       IF #INO_tTrack.rgtTrackMachine[#IN_dMachineIndex].tUserData.dGetDownstreamIndex >= 0 THEN
           #AUX_xValidDwCap := TRUE;
           #OS_xNewCapDw := TRUE;            
           #AUX_dDwCapIndex := #INO_tTrack.rgtTrackMachine[#IN_dMachineIndex].tUserData.dGetDownstreamIndex;
       ELSE
           #AUX_xValidDwCap := FALSE;
           #OS_xNewCapDw := FALSE;            
           #AUX_dDwCapIndex := 0;
       END_IF;

       #INO_tTrack.rgtTrackMachine[#IN_dMachineIndex].tUserData.xGetPosReach := FALSE;

   END_IF;
END_REGION

REGION Network 6: ####_HMI_LOGICS_####
END_REGION

REGION Network 7 (SCL): List of HMI logics
   REGION UpdateDistanceSnaproll

   IF #tHMW.xUpdateDistSnap THEN
       #tHMW.xUpdateDistSnap := FALSE;

       #tHMR.dDistanceFromSnaproll_cmm := #tHMW.dDistanceFromSnaproll_cmm;

   END_IF;

   END_REGION
END_REGION

REGION Network 8: ####_ALARMS_####
END_REGION

REGION Network 9 (SCL): Reset alarms
   IF #IN_xResetAlarms THEN

       #TMP_dwValue := 0;

       SCATTER(IN:=#TMP_dwValue,
               OUT=>#tALM.tF);

       SCATTER(IN:=#TMP_dwValue,
               OUT=>#tALM.tS);

       SCATTER(IN:=#TMP_dwValue,
               OUT=>#tALM.tW);

   END_IF;
END_REGION

REGION Network 10: ####_STATUSES_####
END_REGION

REGION Network 11 (SCL): Calculate alarm statuses
   GATHER(IN:=#tALM.tS,
          OUT=>#TMP_dwValue);

   IF #TMP_dwValue <> 0 THEN
       #ST_xStoppingFaults := TRUE;
   ELSE
       #ST_xStoppingFaults := FALSE;
   END_IF;

   GATHER(IN:=#tALM.tF,
          OUT=>#TMP_dwValue);

   IF #TMP_dwValue <> 0 THEN
       #ST_xFaults := TRUE;
   ELSE
       #ST_xFaults := FALSE;
   END_IF;

   GATHER(IN:=#tALM.tW,
          OUT=>#TMP_dwValue);

   IF #TMP_dwValue <> 0 THEN
       #ST_xWarnings := TRUE;
   ELSE
       #ST_xWarnings := FALSE;
   END_IF;
END_REGION

REGION Network 12 (SCL): Glass break calculation
   #INO_tRibbon.rgtGlassBreakRequest[#IN_dGlassBreakMachineIndex].IN_dDistanceSnaproll_cmm := #tHMR.dDistanceFromSnaproll_cmm;
   #INO_tRibbon.rgtGlassBreakRequest[#IN_dGlassBreakMachineIndex].IN_dDownstreamOffset_cmm := #CONST_DBREAKDOWNOFF_CMM;
   #INO_tRibbon.rgtGlassBreakRequest[#IN_dGlassBreakMachineIndex].IN_dUpstreamOffset_cmm := #CONST_DBREAKUPOFF_CMM;

   IF #INO_tRibbon.rgtGlassBreakRequest[#IN_dGlassBreakMachineIndex].OUT_xDataReady THEN
       #ST_xGlassBreak := #INO_tRibbon.rgtGlassBreakRequest[#IN_dGlassBreakMachineIndex].OUT_xGlassBreak;
   END_IF;

   IF #INO_tRibbon.rgtGlassBreakRequest[#IN_dGlassBreakMachineIndex].OUT_xDataReady OR NOT #INO_tRibbon.rgtGlassBreakRequest[#IN_dGlassBreakMachineIndex].IN_xRequestGlassBreak THEN
       #INO_tRibbon.rgtGlassBreakRequest[#IN_dGlassBreakMachineIndex].OUT_xDataReady := FALSE;
       #INO_tRibbon.rgtGlassBreakRequest[#IN_dGlassBreakMachineIndex].IN_xRequestGlassBreak := TRUE;
   END_IF;
END_REGION

REGION Network 13: ####_PHASES_&_LOGICS_####
END_REGION

REGION Network 14: Plate under bridge
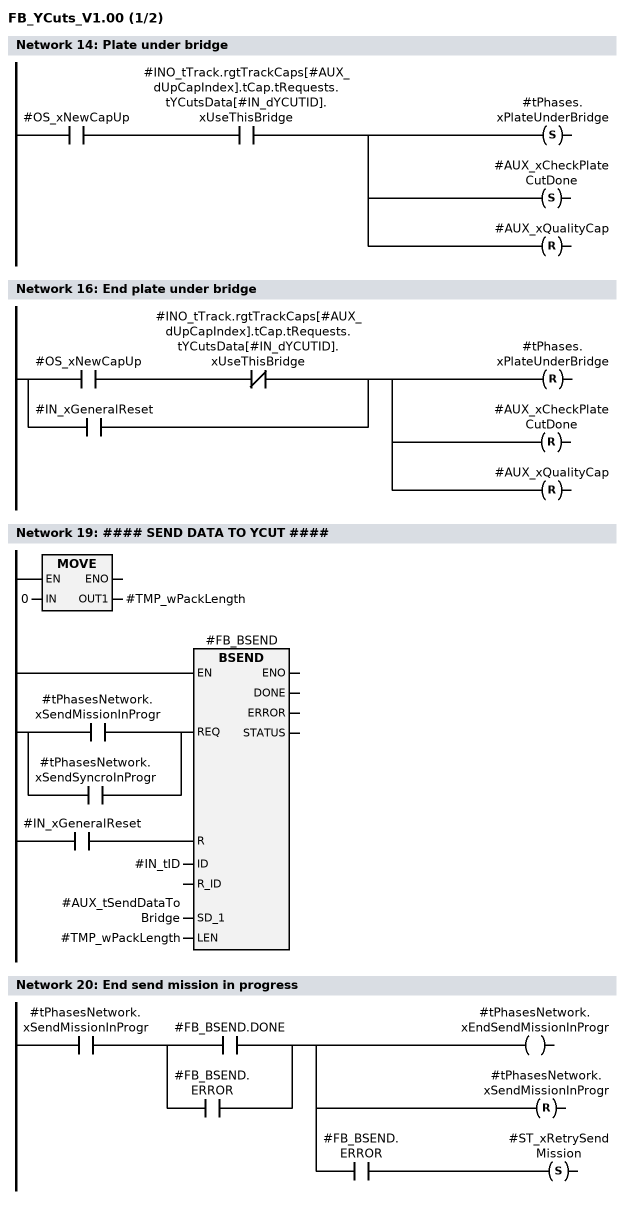
   RUNG wire#powerrail
      Contact( #OS_xNewCapUp )
      Contact( #INO_tTrack.rgtTrackCaps[#AUX_dUpCapIndex].tCap.tRequests.tYCutsData[#IN_dYCUTID].xUseThisBridge )
      wire#w1
      S_Coil( #tPhases.xPlateUnderBridge )
   END_RUNG
   RUNG wire#w1
      S_Coil( #AUX_xCheckPlateCutDone )
   END_RUNG
   RUNG wire#w1
      R_Coil( #AUX_xQualityCap )
   END_RUNG
   // the same network as SCL:
   IF #OS_xNewCapUp AND #INO_tTrack.rgtTrackCaps[#AUX_dUpCapIndex].tCap.tRequests.tYCutsData[#IN_dYCUTID].xUseThisBridge THEN
       #tPhases.xPlateUnderBridge := TRUE;
       #AUX_xCheckPlateCutDone := TRUE;
       #AUX_xQualityCap := FALSE;
   END_IF;
END_REGION

REGION Network 15 (SCL): Tracking plate
   IF #tPhases.xPlateUnderBridge AND #AUX_xValidUpCap AND #AUX_xCheckPlateCutDone  THEN

       IF  #INO_tTrack.rgtTrackCaps[#AUX_dUpCapIndex].tCap.rgtLites[0].dMainDestination = "DQUALITYDESTMASK1" OR
           #INO_tTrack.rgtTrackCaps[#AUX_dUpCapIndex].tCap.rgtLites[0].dMainDestination = "DQUALITYDESTMASK2" OR
           #INO_tTrack.rgtTrackCaps[#AUX_dUpCapIndex].tCap.rgtLites[0].dMainDestination = "DQUALITYDESTMASK3" OR
           #INO_tTrack.rgtTrackCaps[#AUX_dUpCapIndex].tCap.rgtLites[0].dMainDestination = "DQUALITYDESTMASK4" THEN

           IF #INO_tTrack.rgtTrackCaps[#AUX_dUpCapIndex].tCap.tRequests.xYCutSampleTest THEN
               #AUX_xQualityCap := TRUE;
           END_IF;

       END_IF;




       #AUX_dActualRecoverWander_cmm := #INO_tTrack.rgtTrackCaps[#AUX_dUpCapIndex].tCap.dEndCutWander_cmm;

       //Assume that cuts are done
       #INO_tTrack.rgtTrackCaps[#AUX_dUpCapIndex].tCap.tDone.tYCuts[#IN_dYCUTID].rgxHeadsDone := 
                           #INO_tTrack.rgtTrackCaps[#AUX_dUpCapIndex].tCap.tRequests.tYCutsData[#IN_dYCUTID].rgxHeadsRequest;    

       //Evaluate the plate 20% more and 80% less. If missing cut take out the done
       #TMP_dPercLength_cmm := REAL_TO_DINT(DINT_TO_REAL(#INO_tTrack.rgtTrackCaps[#AUX_dUpCapIndex].tCap.dLength_cmm) * 0.2);

       #TMP_dOpenGatePosition_cmm := #TMP_dPercLength_cmm;
       #TMP_dCloseGatePosition_cmm := #INO_tTrack.rgtTrackCaps[#AUX_dUpCapIndex].tCap.dLength_cmm - #TMP_dPercLength_cmm;

       #TMP_dEncOnYCut_cmm := #INO_tEnc.dActualEncoderCounter_cmm + #tHMR.dDistanceFromSnaproll_cmm;

       #TMP_dValue_cmm := #TMP_dEncOnYCut_cmm - #INO_tTrack.rgtTrackCaps[#AUX_dUpCapIndex].tCap.dHeadPositionBTC;   

       #TMP_xRequestIsNotDone := FALSE;

       IF NOT #IN_xSimulationActive   THEN

           IF ((#TMP_dValue_cmm >= #TMP_dOpenGatePosition_cmm) AND (#TMP_dValue_cmm <= #TMP_dCloseGatePosition_cmm)) THEN

               FOR #TMP_dIndex := 0 TO "DMAXYHEADS_IND" DO

                   IF #IN_tIDeviceData.rgxCuttingStatus[#TMP_dIndex] = FALSE AND
                       #INO_tTrack.rgtTrackCaps[#AUX_dUpCapIndex].tCap.tRequests.tYCutsData[#IN_dYCUTID].rgxHeadsRequest[#TMP_dIndex] THEN
                       #INO_tTrack.rgtTrackCaps[#AUX_dUpCapIndex].tCap.tDone.tYCuts[#IN_dYCUTID].rgxHeadsDone[#TMP_dIndex] := FALSE;
                       #TMP_xRequestIsNotDone := TRUE;
                   END_IF;
               END_FOR;
           END_IF;
       END_IF;

       IF #TMP_xRequestIsNotDone THEN

           #AUX_xCheckPlateCutDone := FALSE;

           //Evaluate all the lite. Send to cullet 
           FOR #TMP_dIndex := 0 TO  #INO_tTrack.rgtTrackCaps[#AUX_dUpCapIndex].tCap.dNumLites - 1 DO

               IF #INO_tTrack.rgtTrackCaps[#AUX_dUpCapIndex].tCap.rgtLites[#TMP_dIndex].dMainDestination <> "DCULLETDESTMASK" THEN

                   #INO_tTrack.rgtTrackCaps[#AUX_dUpCapIndex].tCap.rgtLites[#TMP_dIndex].dMainDestination := "DCULLETDESTMASK";
                   #INO_tTrack.rgtTrackCaps[#AUX_dUpCapIndex].tCap.rgtLites[#TMP_dIndex].dAltDestination := 0;
                   #INO_tTrack.rgtTrackCaps[#AUX_dUpCapIndex].tCap.rgtLites[#TMP_dIndex].d2ndDestionation := 0;
                   #INO_tTrack.rgtTrackCaps[#AUX_dUpCapIndex].tCap.rgtLites[#TMP_dIndex].dCulletCause := "DCULLETCAUSE_YCUTMISSING";

               END_IF;
           END_FOR;

           #INO_tTrack.rgtTrackCaps[#AUX_dUpCapIndex].tCap.tRequests.xUpdateDataBPSA := TRUE;
           #INO_tTrack.rgtTrackCaps[#AUX_dUpCapIndex].tCap.tRequests.xUpdateDataBPSB := TRUE;

       END_IF;

   END_IF;
END_REGION

REGION Network 16: End plate under bridge
   RUNG wire#powerrail
      Contact( #OS_xNewCapUp )
      I_Contact( #INO_tTrack.rgtTrackCaps[#AUX_dUpCapIndex].tCap.tRequests.tYCutsData[#IN_dYCUTID].xUseThisBridge )
      wire#w1
      R_Coil( #tPhases.xPlateUnderBridge )
   END_RUNG
   RUNG wire#powerrail
      Contact( #IN_xGeneralReset )
   END_RUNG wire#w1
   RUNG wire#w1
      R_Coil( #AUX_xCheckPlateCutDone )
   END_RUNG
   RUNG wire#w1
      R_Coil( #AUX_xQualityCap )
   END_RUNG
   // the same network as SCL:
   IF (#OS_xNewCapUp AND NOT #INO_tTrack.rgtTrackCaps[#AUX_dUpCapIndex].tCap.tRequests.tYCutsData[#IN_dYCUTID].xUseThisBridge) OR #IN_xGeneralReset THEN
       #tPhases.xPlateUnderBridge := FALSE;
       #AUX_xCheckPlateCutDone := FALSE;
       #AUX_xQualityCap := FALSE;
   END_IF;
END_REGION

REGION Network 17 (SCL): Send mission in progress
   IF NOT #ST_xPhaseInProgressNetwork AND (#INO_tTrack.rgxNewCapAvailable[#IN_dTrackNewCapIndex] OR #ST_xRetrySendMission) AND NOT #IN_xSimulationActive THEN

       #TMP_xTripleEdgeSituation := FALSE;
       #TMP_dOppositeBridgeIndex := 0;
       IF (#INO_tTrack.rgxNewCapAvailable[#IN_dTrackNewCapIndex] AND (NOT #INO_tTrack.tLastPlacedCap.tRequests.tYCutsData[#IN_dYCUTID].xUseThisBridge) 
           AND (#INO_tTrack.tLastPlacedCap.dTEdgeOppOpSide_cmm > 0  OR #INO_tTrack.tLastPlacedCap.dTEdgeOpSide_cmm > 0 )) THEN

           IF #IN_dYCUTID = 1 THEN
               #TMP_dOppositeBridgeIndex := 0;
           ELSE
               #TMP_dOppositeBridgeIndex := 1;
           END_IF;

           IF #INO_tTrack.tLastPlacedCap.tRequests.tYCutsData[#TMP_dOppositeBridgeIndex].xUseThisBridge THEN
             #TMP_xTripleEdgeSituation := TRUE;
           END_IF;
       END_IF;

       IF (#INO_tTrack.rgxNewCapAvailable[#IN_dTrackNewCapIndex] AND #INO_tTrack.tLastPlacedCap.tRequests.tYCutsData[#IN_dYCUTID].xUseThisBridge) OR 
           #TMP_xTripleEdgeSituation  THEN

           #AUX_tSendDataToBridge.tMissionData.dMissionID := #INO_tTrack.tLastPlacedCap.rgtLites[0].dID;
           #AUX_tSendDataToBridge.tMissionData.dMissionStart_cmm := #INO_tTrack.tLastPlacedCap.dHeadPositionBTC - #tHMR.dDistanceFromSnaproll_cmm;
           #AUX_tSendDataToBridge.tMissionData.dMissionEnd_cmm := #INO_tTrack.tLastPlacedCap.dTailPositionBTC - #tHMR.dDistanceFromSnaproll_cmm;


           //If is a quality sample plate reduce the fireon and off of 5cm
           IF #INO_tTrack.tLastPlacedCap.tRequests.xYCutSampleTest THEN
               #AUX_tSendDataToBridge.tMissionData.dMissionStart_cmm += 20000;
               #AUX_tSendDataToBridge.tMissionData.dMissionEnd_cmm -= 20000;
           END_IF;

           #TMP_dwValue := 0;

           SCATTER(IN:=#TMP_dwValue,
                   OUT=>#AUX_tSendDataToBridge.tMissionData.rgxFireRequest);

           FOR #TMP_dIndex := 0 TO "DMAXYHEADS_IND" DO

               #AUX_tSendDataToBridge.tMissionData.rgxFireRequest[#TMP_dIndex] := 
                               #INO_tTrack.tLastPlacedCap.tRequests.tYCutsData[#IN_dYCUTID].rgxHeadsRequest[#TMP_dIndex];

               #AUX_tSendDataToBridge.tMissionData.rgdHeadsPosition_cmm[#TMP_dIndex] :=    
               #INO_tTrack.tLastPlacedCap.tRequests.tYCutsData[#IN_dYCUTID].rgdHeadsPositions[#TMP_dIndex];

               IF #TMP_xTripleEdgeSituation THEN

                   #AUX_tSendDataToBridge.tMissionData.rgdHeadsPosition_cmm[#TMP_dIndex] :=    
                       #INO_tTrack.tLastPlacedCap.tRequests.tYCutsData[#TMP_dOppositeBridgeIndex].rgdHeadsPositions[#TMP_dIndex];

                   IF #TMP_dIndex = #CONST_TRIPLE_FIRSTHEAD AND #INO_tTrack.tLastPlacedCap.dTEdgeOpSide_cmm > 0  THEN
                       #AUX_tSendDataToBridge.tMissionData.rgdHeadsPosition_cmm[#TMP_dIndex]-= #INO_tTrack.tLastPlacedCap.dTEdgeOpSide_cmm;    
                       #AUX_tSendDataToBridge.tMissionData.rgxFireRequest[#TMP_dIndex] := TRUE; 
                   ELSIF #TMP_dIndex = #CONST_TRIPLE_LASTHEAD AND #INO_tTrack.tLastPlacedCap.dTEdgeOppOpSide_cmm > 0  THEN   
                       #AUX_tSendDataToBridge.tMissionData.rgdHeadsPosition_cmm[#TMP_dIndex]+= #INO_tTrack.tLastPlacedCap.dTEdgeOppOpSide_cmm;    
                       #AUX_tSendDataToBridge.tMissionData.rgxFireRequest[#TMP_dIndex] := TRUE; 
                   END_IF;
               END_IF;

           END_FOR;



           #tPhasesNetwork.xSendMissionInProgr := TRUE;
           #ST_xRetrySendMission := FALSE;

           #INO_tTrack.rgxNewCapAvailable[#IN_dTrackNewCapIndex] := FALSE;
       END_IF;

       IF #ST_xRetrySendMission = TRUE THEN
           #tPhasesNetwork.xSendMissionInProgr := TRUE;
           #ST_xRetrySendMission := FALSE;
       END_IF;

       IF #INO_tTrack.rgxNewCapAvailable[#IN_dTrackNewCapIndex] = TRUE THEN
           #INO_tTrack.rgxNewCapAvailable[#IN_dTrackNewCapIndex] := FALSE;
       END_IF;
   END_IF;
END_REGION

REGION Network 18 (SCL): Send data to bridge
   IF NOT #ST_xPhaseInProgressNetwork AND (#INO_tEnc.rgxMetersForYCuts[#IN_dYCUTID] OR #ST_xRetrySendSyncro) THEN

       IF #INO_tEnc.rgxMetersForYCuts[#IN_dYCUTID] THEN

           #AUX_tSendDataToBridge.tSyncroData.dMissionID+= 1;
           #AUX_tSendDataToBridge.tSyncroData.dSynchroValue_cmm := #INO_tEnc.dLastMeterValue_cmm;        

           #INO_tEnc.rgxMetersForYCuts[#IN_dYCUTID] := FALSE;
           #ST_xRetrySendSyncro := FALSE;
           #tPhasesNetwork.xSendSyncroInProgr := TRUE;
       END_IF;

       IF #ST_xRetrySendSyncro THEN
           #ST_xRetrySendSyncro := FALSE;
           #tPhasesNetwork.xSendSyncroInProgr := TRUE;
       END_IF;

   END_IF;
END_REGION

REGION Network 19: #### SEND DATA TO YCUT ####
   #TMP_wPackLength := 0;
   #FB_BSEND(REQ := #tPhasesNetwork.xSendMissionInProgr OR #tPhasesNetwork.xSendSyncroInProgr,   // BSEND
             R := #IN_xGeneralReset,
             ID := #IN_tID,
             SD_1 := #AUX_tSendDataToBridge,
             LEN := #TMP_wPackLength);
END_REGION

REGION Network 20: End send mission in progress
   RUNG wire#powerrail
      Contact( #tPhasesNetwork.xSendMissionInProgr )
      wire#w1
      Contact( #FB_BSEND.DONE )
      wire#w2
      Coil( #tPhasesNetwork.xEndSendMissionInProgr )
   END_RUNG
   RUNG wire#w1
      Contact( #FB_BSEND.ERROR )
   END_RUNG wire#w2
   RUNG wire#w2
      R_Coil( #tPhasesNetwork.xSendMissionInProgr )
   END_RUNG
   RUNG wire#w2
      Contact( #FB_BSEND.ERROR )
      S_Coil( #ST_xRetrySendMission )
   END_RUNG
   // the same network as SCL:
   #tPhasesNetwork.xEndSendMissionInProgr := #tPhasesNetwork.xSendMissionInProgr AND (#FB_BSEND.DONE OR #FB_BSEND.ERROR);
   IF #tPhasesNetwork.xEndSendMissionInProgr THEN #tPhasesNetwork.xSendMissionInProgr := FALSE; END_IF;
   IF #tPhasesNetwork.xEndSendMissionInProgr AND #FB_BSEND.ERROR THEN #ST_xRetrySendMission := TRUE; END_IF;
END_REGION

REGION Network 21: End send syncro in progress
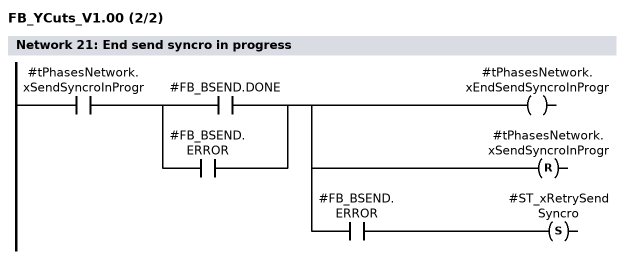
   RUNG wire#powerrail
      Contact( #tPhasesNetwork.xSendSyncroInProgr )
      wire#w1
      Contact( #FB_BSEND.DONE )
      wire#w2
      Coil( #tPhasesNetwork.xEndSendSyncroInProgr )
   END_RUNG
   RUNG wire#w1
      Contact( #FB_BSEND.ERROR )
   END_RUNG wire#w2
   RUNG wire#w2
      R_Coil( #tPhasesNetwork.xSendSyncroInProgr )
   END_RUNG
   RUNG wire#w2
      Contact( #FB_BSEND.ERROR )
      S_Coil( #ST_xRetrySendSyncro )
   END_RUNG
   // the same network as SCL:
   #tPhasesNetwork.xEndSendSyncroInProgr := #tPhasesNetwork.xSendSyncroInProgr AND (#FB_BSEND.DONE OR #FB_BSEND.ERROR);
   IF #tPhasesNetwork.xEndSendSyncroInProgr THEN #tPhasesNetwork.xSendSyncroInProgr := FALSE; END_IF;
   IF #tPhasesNetwork.xEndSendSyncroInProgr AND #FB_BSEND.ERROR THEN #ST_xRetrySendSyncro := TRUE; END_IF;
END_REGION

REGION Network 22 (SCL): Calculare phase in progress
   GATHER(IN:=#tPhases,
          OUT=>#TMP_dwValue);

   IF #TMP_dwValue <> 0 THEN
       #ST_xPhaseInProgress := TRUE;
   ELSE
       #ST_xPhaseInProgress := FALSE;
   END_IF;

   GATHER(IN := #tPhasesNetwork,
           OUT => #TMP_dwValue);

   IF  #TMP_dwValue <> 0 THEN
       #ST_xPhaseInProgressNetwork := TRUE;
   ELSE
       #ST_xPhaseInProgressNetwork := FALSE;
   END_IF;
END_REGION

REGION Network 23: ####_OUTPUT_####
END_REGION

REGION Network 24 (SCL): Compile IDevice output
   #OUT_tIDeviceData.xCycleON := #IN_xCycleON;
   #OUT_tIDeviceData.xGlassBreak := #ST_xGlassBreak;
   #OUT_tIDeviceData.xPLCActive0 := TRUE;
   #OUT_tIDeviceData.xPLCActive1 := FALSE;
   #OUT_tIDeviceData.xQLTplate := #AUX_xQualityCap;
   #OUT_tIDeviceData.xResetAnomaly := #IN_xResetAlarms;
   #OUT_tIDeviceData.xResetBuffers := #IN_xGeneralReset;
END_REGION

REGION Network 25 (SCL): Compile bridge status output
   IF #IN_xSimulationActive THEN

       #OUT_tBridgeStatus.dBridgeStatus := 3;

       #TMP_wValue := W#16#FFFF;

       SCATTER(IN := #TMP_wValue,
               OUT=> #OUT_tBridgeStatus.rgxHeadProdOn);

       IF #OS_xNewCapUp THEN

           //Put to 0 the fire mask
           #TMP_wValue := 0;

           SCATTER(IN:=#TMP_wValue,
                   OUT=>#OUT_tBridgeStatus.rgxFireON);

           IF #INO_tTrack.rgtTrackCaps[#AUX_dUpCapIndex].tCap.tRequests.tYCutsData[#IN_dYCUTID].xUseThisBridge THEN

               #OUT_tBridgeStatus.rgdPosition_cmm := #INO_tTrack.rgtTrackCaps[#AUX_dUpCapIndex].tCap.tRequests.tYCutsData[#IN_dYCUTID].rgdHeadsPositions;
               #OUT_tBridgeStatus.rgxFireON := #INO_tTrack.rgtTrackCaps[#AUX_dUpCapIndex].tCap.tRequests.tYCutsData[#IN_dYCUTID].rgxHeadsRequest;
               #OUT_tBridgeStatus.rgxArmON := #OUT_tBridgeStatus.rgxFireON;

           END_IF;
       END_IF;
   ELSE

       IF #IN_tIDeviceData.rgxStatus[2] THEN
           #OUT_tBridgeStatus.dBridgeStatus := 3;

           IF #IN_tIDeviceData.rgxStatus[0] THEN
               #OUT_tBridgeStatus.dBridgeStatus := 4;
           END_IF;

       ELSE
           #OUT_tBridgeStatus.dBridgeStatus := 1;
       END_IF;

       #OUT_tBridgeStatus.rgdPosition_cmm := #IN_tIDeviceData.rgdHeadsPositions_cmm;
       #OUT_tBridgeStatus.rgxFireON := #IN_tIDeviceData.rgxCuttingStatus;
       #OUT_tBridgeStatus.rgxHeadProdOn := #IN_tIDeviceData.rgxHeadStatus;

   END_IF;
END_REGION
END_FUNCTION_BLOCK

// folder: 03_Programs_Logics/MCC1200/11_SnapRoll

FUNCTION_BLOCK "FB_Snaproll_V1.00"   // FB10, LAD
TITLE = Snaproll machine V1.00
{ S7_Optimized_Access := 'TRUE' }
VERSION : 0.1
   VAR_INPUT
      IN_dMachineIndex : DInt;   // Tracking machine index
      IN_xCycleON : Bool;   // Cycle ON
      IN_xGeneralReset : Bool;   // General reset
      IN_xResetAlarms : Bool;   // Reset alarms
      IN_xFaultsEnabled : Bool;   // Faults enabled
      INPUT : Struct
         xForceUp : Bool;
         xForceDw : Bool;
      END_STRUCT;
   END_VAR
   VAR_OUTPUT
      tOutputs : Struct   // Outputs
         rgxHLCutDoneXC : Array[0.."DMAXXHEADS_IND"] of Bool;   // HL cut done by xc#x
         xRiseSnap : Bool;   // Rise snaproll
         xContrastActivation : Bool;   // Contrast activation
      END_STRUCT;
   END_VAR
   VAR_IN_OUT
      INO_tTrack : "UDT_CapData_Tracking";   // Tracking plate
      INO_tEnc : "UDT_Encoder";   // Encoder data
   END_VAR
   VAR RETAIN
      tHMW : Struct   // HMI Write data
         dOffsetSnap_cmm : DInt;   // Offset rise snap (- Anticipate + Delay) [mm/100] {mm/100|mm|-300|300|O}
         dMaxPlateLenghtEnableContrast_cmm : DInt;   // Maximum plate lenght for contrast enabling [mm/100] {mm/100|mm|1|7000|O}
         dTimeUp_ms : DInt;   // Time snap in up position [ms] {ms|s|0|1|O}
         dReactTime_ms : DInt;   // Snap reaction time [ms] {ms|s|0|1|O}
         xEnDisManComSnap : Bool;   // Enable disable manual command snaroll {x|x|x|x|O}
         tMan : Struct   // Manual commands
            xUp : Bool;   // Snap roll up {x|x|x|x|O}
            xContrastActivation : Bool;   // Contrast activation {x|x|x|x|O}
            xSpare_2 : Bool;
            xSpare_3 : Bool;
            xSpare_4 : Bool;
            xSpare_5 : Bool;
            xSpare_6 : Bool;
            xSpare_7 : Bool;
            xSpare_8 : Bool;
            xSpare_9 : Bool;
            xSpare_10 : Bool;
            xSpare_11 : Bool;
            xSpare_12 : Bool;
            xSpare_13 : Bool;
            xSpare_14 : Bool;
            xSpare_15 : Bool;
         END_STRUCT;
      END_STRUCT;
      tHMR : Struct   // HMI Read data
         dStatus : DInt;   // Status (1=Idle 3=Up 7=Fault) {x|x|x|x|O}
         xManComEnSnap : Bool;   // Manual command enabled snaproll {x|x|x|x|O}
         tManCmd : Struct   // Manual commands feedback
            xUp : Bool;   // Snap roll up feedback {x|x|x|x|O}
            xContrastActivation : Bool;   // Contrast activation feedback {x|x|x|x|O}
            xSpare_2 : Bool;
            xSpare_3 : Bool;
            xSpare_4 : Bool;
            xSpare_5 : Bool;
            xSpare_6 : Bool;
            xSpare_7 : Bool;
            xSpare_8 : Bool;
            xSpare_9 : Bool;
            xSpare_10 : Bool;
            xSpare_11 : Bool;
            xSpare_12 : Bool;
            xSpare_13 : Bool;
            xSpare_14 : Bool;
            xSpare_15 : Bool;
         END_STRUCT;
      END_STRUCT;
   END_VAR
   VAR
      tALM : Struct   // HMI Alarms
         tS : Struct   // Stopping faults
            xSpare_0 : Bool;
            xSpare_1 : Bool;
            xSpare_2 : Bool;
            xSpare_3 : Bool;
            xSpare_4 : Bool;
            xSpare_5 : Bool;
            xSpare_6 : Bool;
            xSpare_7 : Bool;
            xSpare_8 : Bool;
            xSpare_9 : Bool;
            xSpare_10 : Bool;
            xSpare_11 : Bool;
            xSpare_12 : Bool;
            xSpare_13 : Bool;
            xSpare_14 : Bool;
            xSpare_15 : Bool;
            xSpare_16 : Bool;
            xSpare_17 : Bool;
            xSpare_18 : Bool;
            xSpare_19 : Bool;
            xSpare_20 : Bool;
            xSpare_21 : Bool;
            xSpare_22 : Bool;
            xSpare_23 : Bool;
            xSpare_24 : Bool;
            xSpare_25 : Bool;
            xSpare_26 : Bool;
            xSpare_27 : Bool;
            xSpare_28 : Bool;
            xSpare_29 : Bool;
            xSpare_30 : Bool;
            xSpare_31 : Bool;
         END_STRUCT;
         tF : Struct   // Faults
            xSpare_0 : Bool;
            xSpare_1 : Bool;
            xSpare_2 : Bool;
            xSpare_3 : Bool;
            xSpare_4 : Bool;
            xSpare_5 : Bool;
            xSpare_6 : Bool;
            xSpare_7 : Bool;
            xSpare_8 : Bool;
            xSpare_9 : Bool;
            xSpare_10 : Bool;
            xSpare_11 : Bool;
            xSpare_12 : Bool;
            xSpare_13 : Bool;
            xSpare_14 : Bool;
            xSpare_15 : Bool;
            xSpare_16 : Bool;
            xSpare_17 : Bool;
            xSpare_18 : Bool;
            xSpare_19 : Bool;
            xSpare_20 : Bool;
            xSpare_21 : Bool;
            xSpare_22 : Bool;
            xSpare_23 : Bool;
            xSpare_24 : Bool;
            xSpare_25 : Bool;
            xSpare_26 : Bool;
            xSpare_27 : Bool;
            xSpare_28 : Bool;
            xSpare_29 : Bool;
            xSpare_30 : Bool;
            xSpare_31 : Bool;
         END_STRUCT;
         tW : Struct   // Warnings
            xSpare_0 : Bool;
            xSpare_1 : Bool;
            xSpare_2 : Bool;
            xSpare_3 : Bool;
            xSpare_4 : Bool;
            xSpare_5 : Bool;
            xSpare_6 : Bool;
            xSpare_7 : Bool;
            xSpare_8 : Bool;
            xSpare_9 : Bool;
            xSpare_10 : Bool;
            xSpare_11 : Bool;
            xSpare_12 : Bool;
            xSpare_13 : Bool;
            xSpare_14 : Bool;
            xSpare_15 : Bool;
            xSpare_16 : Bool;
            xSpare_17 : Bool;
            xSpare_18 : Bool;
            xSpare_19 : Bool;
            xSpare_20 : Bool;
            xSpare_21 : Bool;
            xSpare_22 : Bool;
            xSpare_23 : Bool;
            xSpare_24 : Bool;
            xSpare_25 : Bool;
            xSpare_26 : Bool;
            xSpare_27 : Bool;
            xSpare_28 : Bool;
            xSpare_29 : Bool;
            xSpare_30 : Bool;
            xSpare_31 : Bool;
         END_STRUCT;
      END_STRUCT;
      ST_xPhaseInProgress : Bool;   // Phases are in progress
      AUX_xValidUpCap : Bool;   // Upstream cap is valid
      AUX_xValidDwCap : Bool;   // Downstream cap is valid
      AUX_dUpCapIndex : DInt;   // Index of the upstream cap
      AUX_dDwCapIndex : DInt;   // Index of the downstream cap
      OS_xNewCapUp : Bool;   // New cap arrived upstream
      OS_xNewCapDw : Bool;   // New cap arrived downstream
      OS_xNewCap : Bool;   // New cap arrived
      ST_xStoppingFaults : Bool;   // Stopping faults
      ST_xFaults : Bool;   // Faults
      ST_xWarnings : Bool;   // Warnings
      ST_xOutputEnabled : Bool;   // Output enabled
      ST_xGlassBreak : Bool;   // Glass break under bridge
      AUX_xUpIsQuality : Bool;   // Upstream cap is a quality cap
      AUX_xDwIsQuality : Bool;   // Downstream cap is a quality cap
      AUX_xHLCutDoneActive : Bool;   // Lamp active xcut done
      tPhases : Struct   // Phases
         xRiseSnapUp : Bool;   // Rise snap
         xEndRiseSnapUp : Bool;   // End rise snap
         xContrastDown : Bool;   // Contrast activation
         xEndContrastDown : Bool;   // End contrast activation
         xSpare4 : Bool;
         xSpare5 : Bool;
         xSpare6 : Bool;
         xSpare7 : Bool;
         xSpare8 : Bool;
         xSpare9 : Bool;
         xSpare10 : Bool;
         xSpare11 : Bool;
         xSpare12 : Bool;
         xSpare13 : Bool;
         xSpare14 : Bool;
         xSpare15 : Bool;
         xSpare16 : Bool;
         xSpare17 : Bool;
         xSpare18 : Bool;
         xSpare19 : Bool;
         xSpare20 : Bool;
         xSpare21 : Bool;
         xSpare22 : Bool;
         xSpare23 : Bool;
         xSpare24 : Bool;
         xSpare25 : Bool;
         xSpare26 : Bool;
         xSpare27 : Bool;
         xSpare28 : Bool;
         xSpare29 : Bool;
         xSpare30 : Bool;
         xSpare31 : Bool;
      END_STRUCT;
      tmON_ContrastDownElaps : "UDT_IECTON_V1.00";   // TimeON contrast down elapsed time
      tmON_RiseUpSnapElaps : "UDT_IECTON_V1.00";   // TimeON snap up elapsed time
      tmON_LampCutDone : "UDT_IECTON_V1.00";   // Delay off lamp Cut Done
      ST_xOuputEnable : Bool;   // Output enabled
   END_VAR
   VAR_TEMP
      TMP_dwValue : DWord;
      TMP_xCompileMissionData : Bool;
      TMP_dIndex : DInt;
      TMP_wPackLength : Word;
      TMP_xRetrySendMissionWithNewMission : Bool;
      TMP_xRetrySendSyncroWithNewSyncro : Bool;
      TMP_xCompileSyncroData : Bool;
      TMP_xNewCapAvailable : Bool;
      ST_xCondOkManSnap : Bool;   // Condition ok manual command snap
      TMP_wValue : Word;
      TMP_dValue : DInt;
   END_VAR
   VAR CONSTANT
      CONST_DSTATUS_IDLE : DInt := 1;   // Status idle
      CONST_DSTATUS_UP : DInt := 3;   // Status up
      CONST_DSTATUS_ANOMALY : DInt := 7;   // Status anomaly
      CONST_DLIMIT_USESNAP_CMM : DInt := 30100;   // Limit to use snap roll [mm/100]
      CONST_DIST_CONTRASTFROMSNAP : Real := 30000.0;   // Distance from contrast to snaproll [mm/100]
   END_VAR
BEGIN

REGION Network 1: ####_CONSTANTS_####
END_REGION

REGION Network 2: ####_MATCH_####
END_REGION

REGION Network 3 (SCL): Move data information to tracking
   #INO_tTrack.rgtTrackMachine[#IN_dMachineIndex].tUserData.dSetDistanceSnap_cmm := (#tHMW.dOffsetSnap_cmm)*-1;
   #INO_tTrack.rgtTrackMachine[#IN_dMachineIndex].tUserData.dSetMachReacTime_ms := #tHMW.dReactTime_ms;
END_REGION

REGION Network 4 (SCL): Manage tracking call

   #OS_xNewCapUp := FALSE;
   #OS_xNewCapDw := FALSE;
   #OS_xNewCap := FALSE;

   IF #INO_tTrack.rgtTrackMachine[#IN_dMachineIndex].tUserData.xGetPosReach THEN

       IF (NOT #ST_xPhaseInProgress) THEN

           #OS_xNewCap := TRUE;

           IF #INO_tTrack.rgtTrackMachine[#IN_dMachineIndex].tUserData.dGetUpstremIndex >= 0 THEN
               #AUX_xValidUpCap := TRUE;
               #OS_xNewCapUp := TRUE;            
               #AUX_dUpCapIndex := #INO_tTrack.rgtTrackMachine[#IN_dMachineIndex].tUserData.dGetUpstremIndex;
           ELSE
               #AUX_xValidUpCap := FALSE;
               #OS_xNewCapUp := FALSE;            
               #AUX_dUpCapIndex := 0;
           END_IF;

           IF #INO_tTrack.rgtTrackMachine[#IN_dMachineIndex].tUserData.dGetDownstreamIndex >= 0 THEN
               #AUX_xValidDwCap := TRUE;
               #OS_xNewCapDw := TRUE;            
               #AUX_dDwCapIndex := #INO_tTrack.rgtTrackMachine[#IN_dMachineIndex].tUserData.dGetDownstreamIndex;
           ELSE
               #AUX_xValidDwCap := FALSE;
               #OS_xNewCapDw := FALSE;            
               #AUX_dDwCapIndex := 0;
           END_IF;



       END_IF;

       #INO_tTrack.rgtTrackMachine[#IN_dMachineIndex].tUserData.xGetPosReach := FALSE;

   END_IF;
END_REGION

REGION Network 5: ####_HMI_LOGICS_####
END_REGION

REGION Network 6 (SCL): List of HMI logics
END_REGION

REGION Network 7: Condition ok manual command
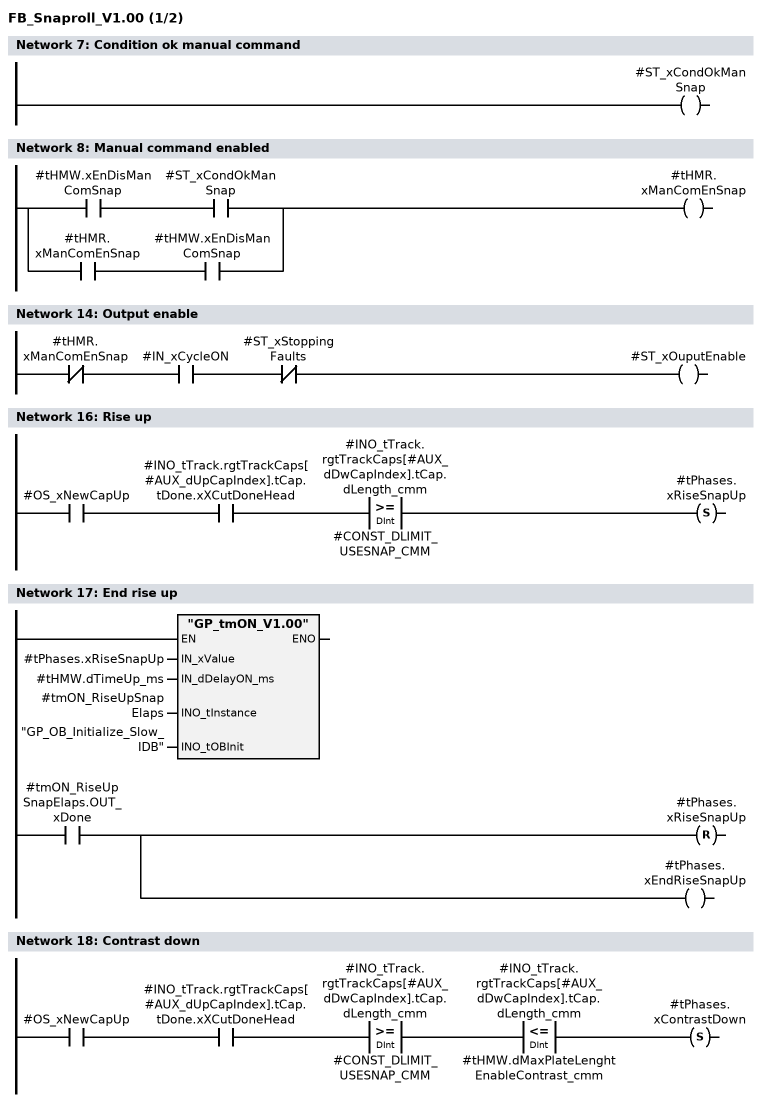
   RUNG wire#powerrail
      Coil( #ST_xCondOkManSnap )
   END_RUNG
   // the same network as SCL:
   #ST_xCondOkManSnap := TRUE;
END_REGION

REGION Network 8: Manual command enabled
   RUNG wire#powerrail
      Contact( #tHMW.xEnDisManComSnap )
      Contact( #ST_xCondOkManSnap )
      wire#w1
      Coil( #tHMR.xManComEnSnap )
   END_RUNG
   RUNG wire#powerrail
      Contact( #tHMR.xManComEnSnap )
      Contact( #tHMW.xEnDisManComSnap )
   END_RUNG wire#w1
   // the same network as SCL:
   #tHMR.xManComEnSnap := (#tHMW.xEnDisManComSnap AND #ST_xCondOkManSnap) OR (#tHMR.xManComEnSnap AND #tHMW.xEnDisManComSnap);
END_REGION

REGION Network 9: ####_ALARMS_####
END_REGION

REGION Network 10 (SCL): Reset alarms
   IF #IN_xResetAlarms THEN

       #TMP_dwValue := 0;

       SCATTER(IN:=#TMP_dwValue,
               OUT=>#tALM.tF);

       SCATTER(IN:=#TMP_dwValue,
               OUT=>#tALM.tS);

       SCATTER(IN:=#TMP_dwValue,
               OUT=>#tALM.tW);

   END_IF;
END_REGION

REGION Network 11: ####_STATUSES_####
END_REGION

REGION Network 12 (SCL): Calculate alarm statuses
   GATHER(IN:=#tALM.tS,
          OUT=>#TMP_dwValue);

   IF #TMP_dwValue <> 0 THEN
       #ST_xStoppingFaults := TRUE;
   ELSE
       #ST_xStoppingFaults := FALSE;
   END_IF;

   GATHER(IN:=#tALM.tF,
          OUT=>#TMP_dwValue);

   IF #TMP_dwValue <> 0 THEN
       #ST_xFaults := TRUE;
   ELSE
       #ST_xFaults := FALSE;
   END_IF;

   GATHER(IN:=#tALM.tW,
          OUT=>#TMP_dwValue);

   IF #TMP_dwValue <> 0 THEN
       #ST_xWarnings := TRUE;
   ELSE
       #ST_xWarnings := FALSE;
   END_IF;
END_REGION

REGION Network 13 (SCL): Reset manual commands
   IF NOT #tHMR.xManComEnSnap THEN

       #TMP_wValue := 0;

       SCATTER(IN:=#TMP_wValue,
               OUT=>#tHMW.tMan);

   END_IF;
END_REGION

REGION Network 14: Output enable
   RUNG wire#powerrail
      I_Contact( #tHMR.xManComEnSnap )
      Contact( #IN_xCycleON )
      I_Contact( #ST_xStoppingFaults )
      Coil( #ST_xOuputEnable )
   END_RUNG
   // the same network as SCL:
   #ST_xOuputEnable := NOT #tHMR.xManComEnSnap AND #IN_xCycleON AND NOT #ST_xStoppingFaults;
END_REGION

REGION Network 15: ####_PHASES_&_LOGICS_####
END_REGION

REGION Network 16: Rise up
   RUNG wire#powerrail
      Contact( #OS_xNewCapUp )
      Contact( #INO_tTrack.rgtTrackCaps[#AUX_dUpCapIndex].tCap.tDone.xXCutDoneHead )
      { S7_Templates := "SrcType := DInt" } GE_Contact(in1 := #INO_tTrack.rgtTrackCaps[#AUX_dDwCapIndex].tCap.dLength_cmm, in2 := #CONST_DLIMIT_USESNAP_CMM)
      S_Coil( #tPhases.xRiseSnapUp )
   END_RUNG
   // the same network as SCL:
   IF #OS_xNewCapUp AND #INO_tTrack.rgtTrackCaps[#AUX_dUpCapIndex].tCap.tDone.xXCutDoneHead AND (#INO_tTrack.rgtTrackCaps[#AUX_dDwCapIndex].tCap.dLength_cmm >= #CONST_DLIMIT_USESNAP_CMM) THEN
       #tPhases.xRiseSnapUp := TRUE;
   END_IF;
END_REGION

REGION Network 17: End rise up
   RUNG wire#powerrail
      "GP_tmON_V1.00"(IN_xValue := #tPhases.xRiseSnapUp, IN_dDelayON_ms := #tHMW.dTimeUp_ms, INO_tInstance := #tmON_RiseUpSnapElaps, INO_tOBInit := "GP_OB_Initialize_Slow_IDB")
   END_RUNG
   RUNG wire#powerrail
      Contact( #tmON_RiseUpSnapElaps.OUT_xDone )
      wire#w1
      R_Coil( #tPhases.xRiseSnapUp )
   END_RUNG
   RUNG wire#w1
      Coil( #tPhases.xEndRiseSnapUp )
   END_RUNG
   // the same network as SCL:
   "GP_tmON_V1.00"(IN_xValue := #tPhases.xRiseSnapUp,
                   IN_dDelayON_ms := #tHMW.dTimeUp_ms,
                   INO_tInstance := #tmON_RiseUpSnapElaps,
                   INO_tOBInit := "GP_OB_Initialize_Slow_IDB");
   IF #tmON_RiseUpSnapElaps.OUT_xDone THEN #tPhases.xRiseSnapUp := FALSE; END_IF;
   #tPhases.xEndRiseSnapUp := #tmON_RiseUpSnapElaps.OUT_xDone;
END_REGION
